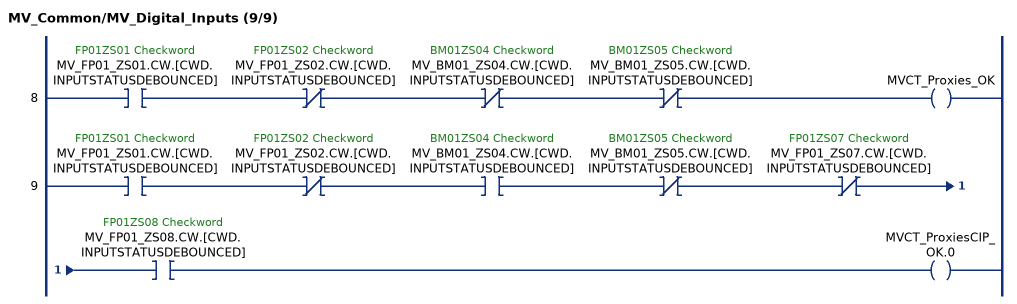
   8: XIC(MV_FP01_ZS01.CW.[CWD.INPUTSTATUSDEBOUNCED])XIO(MV_FP01_ZS02.CW.[CWD.INPUTSTATUSDEBOUNCED])XIO(MV_BM01_ZS04.CW.[CWD.INPUTSTATUSDEBOUNCED])XIO(MV_BM01_ZS05.CW.[CWD.INPUTSTATUSDEBOUNCED])OTE(MVCT_Proxies_OK);
   9: XIC(MV_FP01_ZS01.CW.[CWD.INPUTSTATUSDEBOUNCED])XIO(MV_FP01_ZS02.CW.[CWD.INPUTSTATUSDEBOUNCED])XIC(MV_BM01_ZS04.CW.[CWD.INPUTSTATUSDEBOUNCED])XIO(MV_BM01_ZS05.CW.[CWD.INPUTSTATUSDEBOUNCED])XIO(MV_FP01_ZS07.CW.[CWD.INPUTSTATUSDEBOUNCED])XIC(MV_FP01_ZS08.CW.[CWD.INPUTSTATUSDEBOUNCED])OTE(MVCT_ProxiesCIP_OK.0);
END_ROUTINE

ROUTINE MV_Digital_Outputs   (* ladder *)
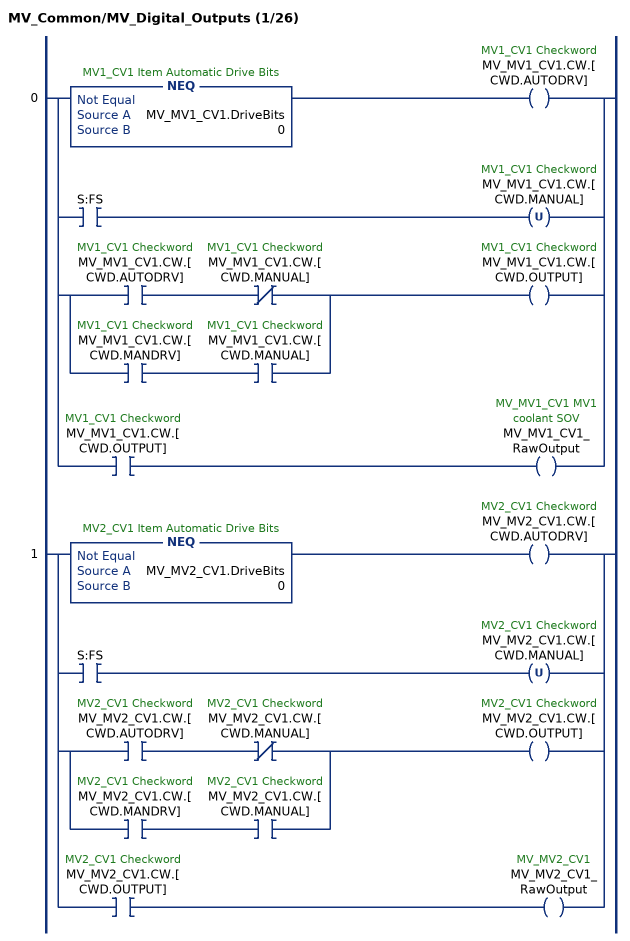
   0: [NEQ(MV_MV1_CV1.DriveBits,0) OTE(MV_MV1_CV1.CW.[CWD.AUTODRV]) ,XIC(S:FS) OTU(MV_MV1_CV1.CW.[CWD.MANUAL]) ,[XIC(MV_MV1_CV1.CW.[CWD.AUTODRV]) XIO(MV_MV1_CV1.CW.[CWD.MANUAL]) ,XIC(MV_MV1_CV1.CW.[CWD.MANDRV]) XIC(MV_MV1_CV1.CW.[CWD.MANUAL]) ] OTE(MV_MV1_CV1.CW.[CWD.OUTPUT]) ,XIC(MV_MV1_CV1.CW.[CWD.OUTPUT]) OTE(MV_MV1_CV1_RawOutput) ];
   1: [NEQ(MV_MV2_CV1.DriveBits,0) OTE(MV_MV2_CV1.CW.[CWD.AUTODRV]) ,XIC(S:FS) OTU(MV_MV2_CV1.CW.[CWD.MANUAL]) ,[XIC(MV_MV2_CV1.CW.[CWD.AUTODRV]) XIO(MV_MV2_CV1.CW.[CWD.MANUAL]) ,XIC(MV_MV2_CV1.CW.[CWD.MANDRV]) XIC(MV_MV2_CV1.CW.[CWD.MANUAL]) ] OTE(MV_MV2_CV1.CW.[CWD.OUTPUT]) ,XIC(MV_MV2_CV1.CW.[CWD.OUTPUT]) OTE(MV_MV2_CV1_RawOutput) ];
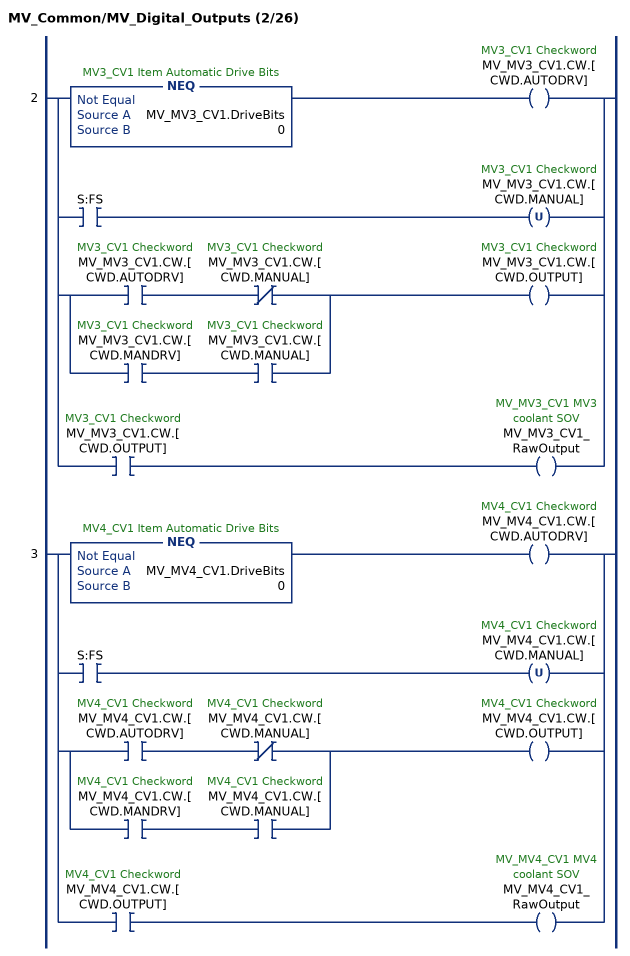
   2: [NEQ(MV_MV3_CV1.DriveBits,0) OTE(MV_MV3_CV1.CW.[CWD.AUTODRV]) ,XIC(S:FS) OTU(MV_MV3_CV1.CW.[CWD.MANUAL]) ,[XIC(MV_MV3_CV1.CW.[CWD.AUTODRV]) XIO(MV_MV3_CV1.CW.[CWD.MANUAL]) ,XIC(MV_MV3_CV1.CW.[CWD.MANDRV]) XIC(MV_MV3_CV1.CW.[CWD.MANUAL]) ] OTE(MV_MV3_CV1.CW.[CWD.OUTPUT]) ,XIC(MV_MV3_CV1.CW.[CWD.OUTPUT]) OTE(MV_MV3_CV1_RawOutput) ];
   3: [NEQ(MV_MV4_CV1.DriveBits,0) OTE(MV_MV4_CV1.CW.[CWD.AUTODRV]) ,XIC(S:FS) OTU(MV_MV4_CV1.CW.[CWD.MANUAL]) ,[XIC(MV_MV4_CV1.CW.[CWD.AUTODRV]) XIO(MV_MV4_CV1.CW.[CWD.MANUAL]) ,XIC(MV_MV4_CV1.CW.[CWD.MANDRV]) XIC(MV_MV4_CV1.CW.[CWD.MANUAL]) ] OTE(MV_MV4_CV1.CW.[CWD.OUTPUT]) ,XIC(MV_MV4_CV1.CW.[CWD.OUTPUT]) OTE(MV_MV4_CV1_RawOutput) ];
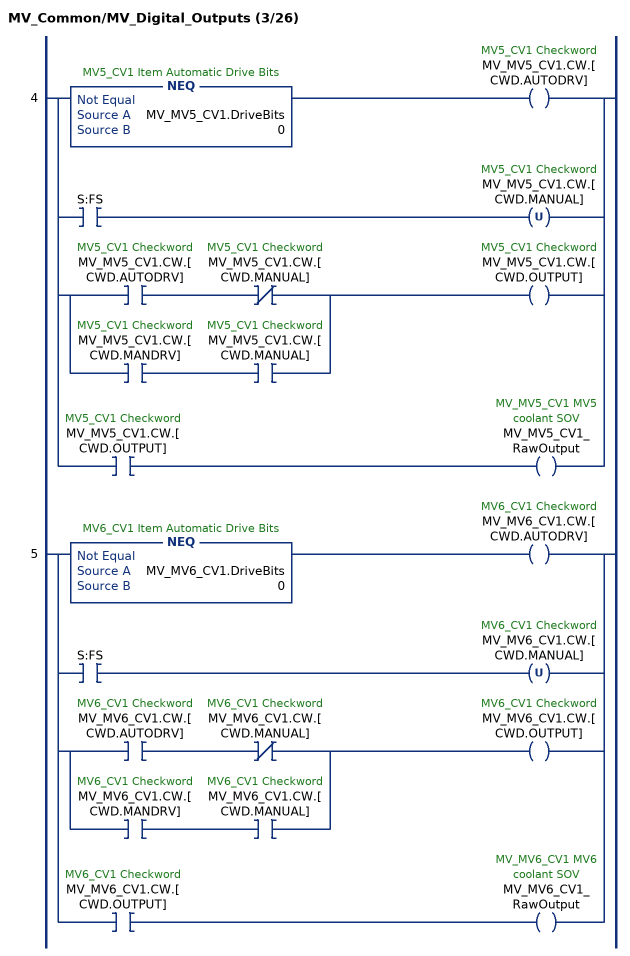
   4: [NEQ(MV_MV5_CV1.DriveBits,0) OTE(MV_MV5_CV1.CW.[CWD.AUTODRV]) ,XIC(S:FS) OTU(MV_MV5_CV1.CW.[CWD.MANUAL]) ,[XIC(MV_MV5_CV1.CW.[CWD.AUTODRV]) XIO(MV_MV5_CV1.CW.[CWD.MANUAL]) ,XIC(MV_MV5_CV1.CW.[CWD.MANDRV]) XIC(MV_MV5_CV1.CW.[CWD.MANUAL]) ] OTE(MV_MV5_CV1.CW.[CWD.OUTPUT]) ,XIC(MV_MV5_CV1.CW.[CWD.OUTPUT]) OTE(MV_MV5_CV1_RawOutput) ];
   5: [NEQ(MV_MV6_CV1.DriveBits,0) OTE(MV_MV6_CV1.CW.[CWD.AUTODRV]) ,XIC(S:FS) OTU(MV_MV6_CV1.CW.[CWD.MANUAL]) ,[XIC(MV_MV6_CV1.CW.[CWD.AUTODRV]) XIO(MV_MV6_CV1.CW.[CWD.MANUAL]) ,XIC(MV_MV6_CV1.CW.[CWD.MANDRV]) XIC(MV_MV6_CV1.CW.[CWD.MANUAL]) ] OTE(MV_MV6_CV1.CW.[CWD.OUTPUT]) ,XIC(MV_MV6_CV1.CW.[CWD.OUTPUT]) OTE(MV_MV6_CV1_RawOutput) ];
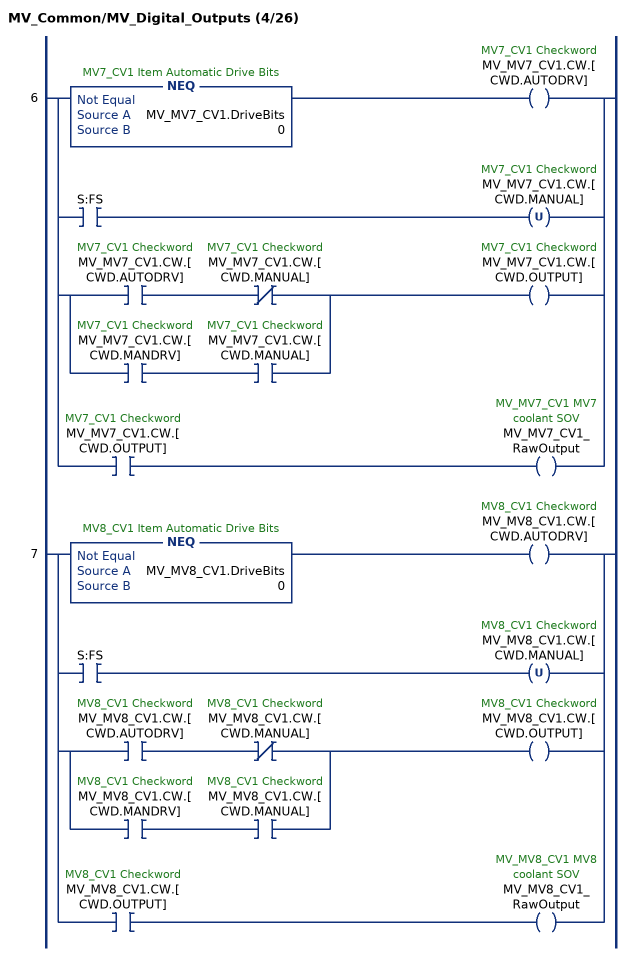
   6: [NEQ(MV_MV7_CV1.DriveBits,0) OTE(MV_MV7_CV1.CW.[CWD.AUTODRV]) ,XIC(S:FS) OTU(MV_MV7_CV1.CW.[CWD.MANUAL]) ,[XIC(MV_MV7_CV1.CW.[CWD.AUTODRV]) XIO(MV_MV7_CV1.CW.[CWD.MANUAL]) ,XIC(MV_MV7_CV1.CW.[CWD.MANDRV]) XIC(MV_MV7_CV1.CW.[CWD.MANUAL]) ] OTE(MV_MV7_CV1.CW.[CWD.OUTPUT]) ,XIC(MV_MV7_CV1.CW.[CWD.OUTPUT]) OTE(MV_MV7_CV1_RawOutput) ];
   7: [NEQ(MV_MV8_CV1.DriveBits,0) OTE(MV_MV8_CV1.CW.[CWD.AUTODRV]) ,XIC(S:FS) OTU(MV_MV8_CV1.CW.[CWD.MANUAL]) ,[XIC(MV_MV8_CV1.CW.[CWD.AUTODRV]) XIO(MV_MV8_CV1.CW.[CWD.MANUAL]) ,XIC(MV_MV8_CV1.CW.[CWD.MANDRV]) XIC(MV_MV8_CV1.CW.[CWD.MANUAL]) ] OTE(MV_MV8_CV1.CW.[CWD.OUTPUT]) ,XIC(MV_MV8_CV1.CW.[CWD.OUTPUT]) OTE(MV_MV8_CV1_RawOutput) ];
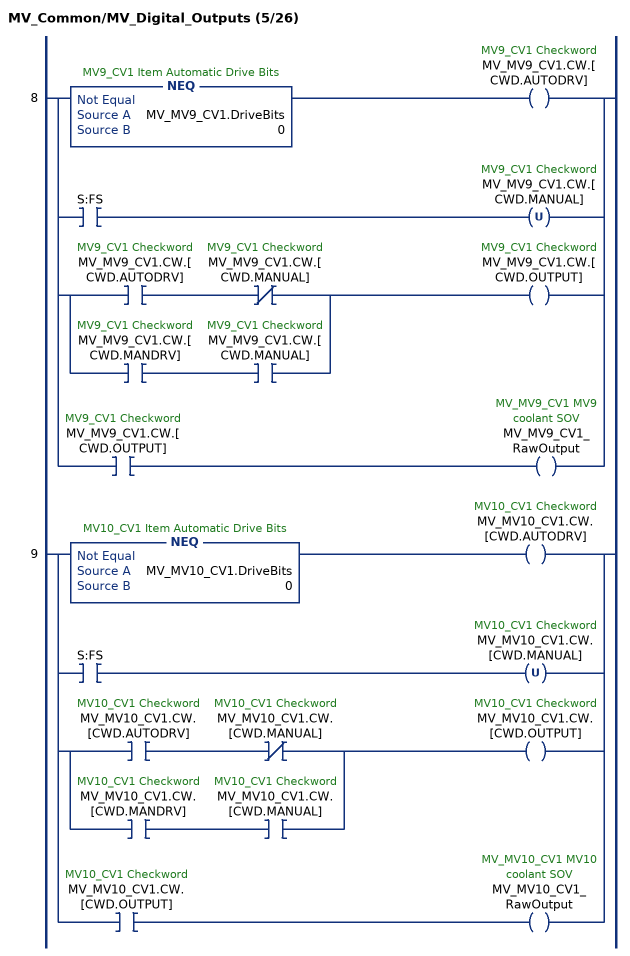
   8: [NEQ(MV_MV9_CV1.DriveBits,0) OTE(MV_MV9_CV1.CW.[CWD.AUTODRV]) ,XIC(S:FS) OTU(MV_MV9_CV1.CW.[CWD.MANUAL]) ,[XIC(MV_MV9_CV1.CW.[CWD.AUTODRV]) XIO(MV_MV9_CV1.CW.[CWD.MANUAL]) ,XIC(MV_MV9_CV1.CW.[CWD.MANDRV]) XIC(MV_MV9_CV1.CW.[CWD.MANUAL]) ] OTE(MV_MV9_CV1.CW.[CWD.OUTPUT]) ,XIC(MV_MV9_CV1.CW.[CWD.OUTPUT]) OTE(MV_MV9_CV1_RawOutput) ];
   9: [NEQ(MV_MV10_CV1.DriveBits,0) OTE(MV_MV10_CV1.CW.[CWD.AUTODRV]) ,XIC(S:FS) OTU(MV_MV10_CV1.CW.[CWD.MANUAL]) ,[XIC(MV_MV10_CV1.CW.[CWD.AUTODRV]) XIO(MV_MV10_CV1.CW.[CWD.MANUAL]) ,XIC(MV_MV10_CV1.CW.[CWD.MANDRV]) XIC(MV_MV10_CV1.CW.[CWD.MANUAL]) ] OTE(MV_MV10_CV1.CW.[CWD.OUTPUT]) ,XIC(MV_MV10_CV1.CW.[CWD.OUTPUT]) OTE(MV_MV10_CV1_RawOutput) ];
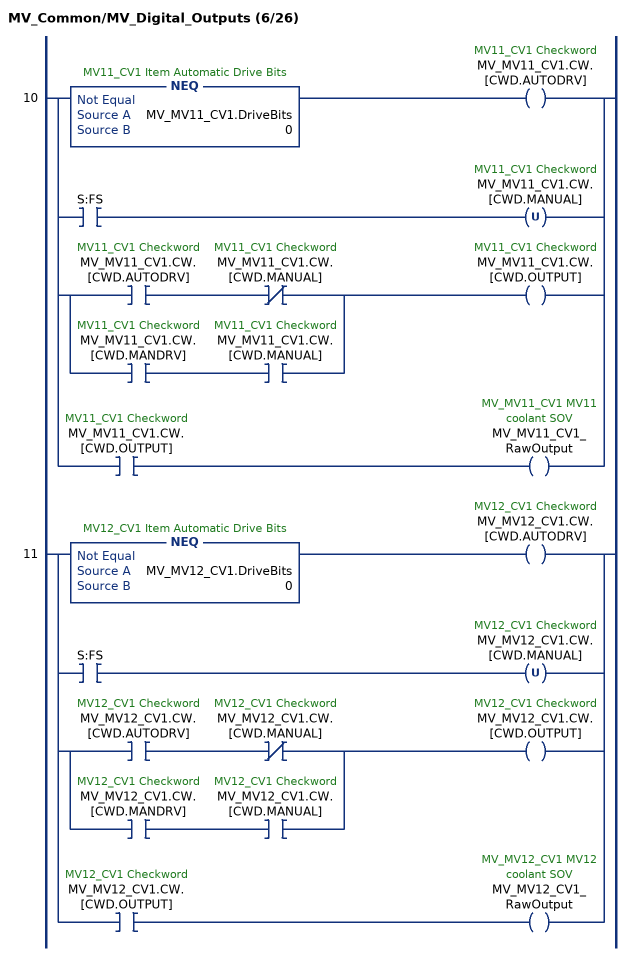
   10: [NEQ(MV_MV11_CV1.DriveBits,0) OTE(MV_MV11_CV1.CW.[CWD.AUTODRV]) ,XIC(S:FS) OTU(MV_MV11_CV1.CW.[CWD.MANUAL]) ,[XIC(MV_MV11_CV1.CW.[CWD.AUTODRV]) XIO(MV_MV11_CV1.CW.[CWD.MANUAL]) ,XIC(MV_MV11_CV1.CW.[CWD.MANDRV]) XIC(MV_MV11_CV1.CW.[CWD.MANUAL]) ] OTE(MV_MV11_CV1.CW.[CWD.OUTPUT]) ,XIC(MV_MV11_CV1.CW.[CWD.OUTPUT]) OTE(MV_MV11_CV1_RawOutput) ];
   11: [NEQ(MV_MV12_CV1.DriveBits,0) OTE(MV_MV12_CV1.CW.[CWD.AUTODRV]) ,XIC(S:FS) OTU(MV_MV12_CV1.CW.[CWD.MANUAL]) ,[XIC(MV_MV12_CV1.CW.[CWD.AUTODRV]) XIO(MV_MV12_CV1.CW.[CWD.MANUAL]) ,XIC(MV_MV12_CV1.CW.[CWD.MANDRV]) XIC(MV_MV12_CV1.CW.[CWD.MANUAL]) ] OTE(MV_MV12_CV1.CW.[CWD.OUTPUT]) ,XIC(MV_MV12_CV1.CW.[CWD.OUTPUT]) OTE(MV_MV12_CV1_RawOutput) ];
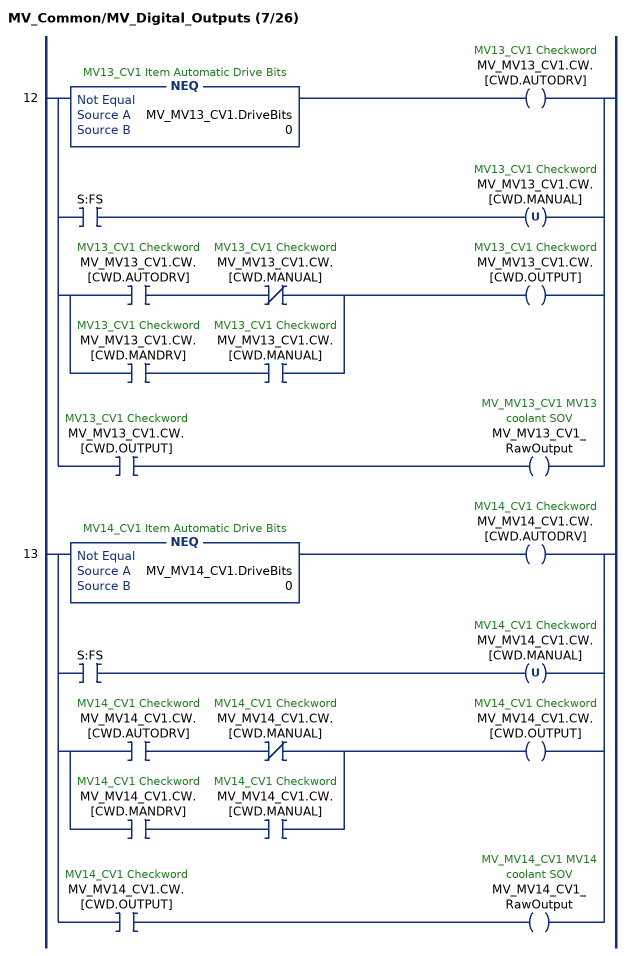
   12: [NEQ(MV_MV13_CV1.DriveBits,0) OTE(MV_MV13_CV1.CW.[CWD.AUTODRV]) ,XIC(S:FS) OTU(MV_MV13_CV1.CW.[CWD.MANUAL]) ,[XIC(MV_MV13_CV1.CW.[CWD.AUTODRV]) XIO(MV_MV13_CV1.CW.[CWD.MANUAL]) ,XIC(MV_MV13_CV1.CW.[CWD.MANDRV]) XIC(MV_MV13_CV1.CW.[CWD.MANUAL]) ] OTE(MV_MV13_CV1.CW.[CWD.OUTPUT]) ,XIC(MV_MV13_CV1.CW.[CWD.OUTPUT]) OTE(MV_MV13_CV1_RawOutput) ];
   13: [NEQ(MV_MV14_CV1.DriveBits,0) OTE(MV_MV14_CV1.CW.[CWD.AUTODRV]) ,XIC(S:FS) OTU(MV_MV14_CV1.CW.[CWD.MANUAL]) ,[XIC(MV_MV14_CV1.CW.[CWD.AUTODRV]) XIO(MV_MV14_CV1.CW.[CWD.MANUAL]) ,XIC(MV_MV14_CV1.CW.[CWD.MANDRV]) XIC(MV_MV14_CV1.CW.[CWD.MANUAL]) ] OTE(MV_MV14_CV1.CW.[CWD.OUTPUT]) ,XIC(MV_MV14_CV1.CW.[CWD.OUTPUT]) OTE(MV_MV14_CV1_RawOutput) ];
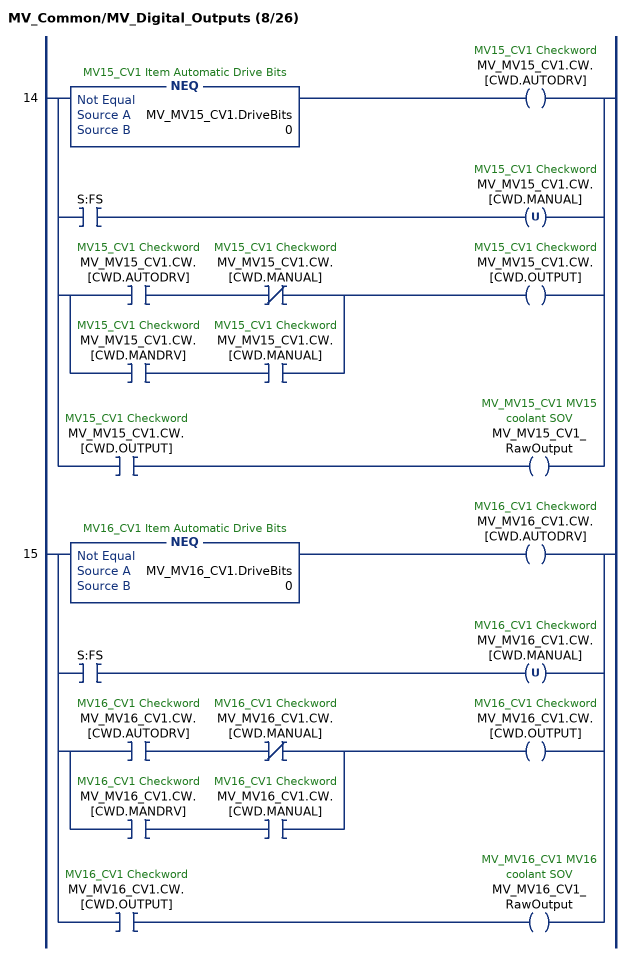
   14: [NEQ(MV_MV15_CV1.DriveBits,0) OTE(MV_MV15_CV1.CW.[CWD.AUTODRV]) ,XIC(S:FS) OTU(MV_MV15_CV1.CW.[CWD.MANUAL]) ,[XIC(MV_MV15_CV1.CW.[CWD.AUTODRV]) XIO(MV_MV15_CV1.CW.[CWD.MANUAL]) ,XIC(MV_MV15_CV1.CW.[CWD.MANDRV]) XIC(MV_MV15_CV1.CW.[CWD.MANUAL]) ] OTE(MV_MV15_CV1.CW.[CWD.OUTPUT]) ,XIC(MV_MV15_CV1.CW.[CWD.OUTPUT]) OTE(MV_MV15_CV1_RawOutput) ];
   15: [NEQ(MV_MV16_CV1.DriveBits,0) OTE(MV_MV16_CV1.CW.[CWD.AUTODRV]) ,XIC(S:FS) OTU(MV_MV16_CV1.CW.[CWD.MANUAL]) ,[XIC(MV_MV16_CV1.CW.[CWD.AUTODRV]) XIO(MV_MV16_CV1.CW.[CWD.MANUAL]) ,XIC(MV_MV16_CV1.CW.[CWD.MANDRV]) XIC(MV_MV16_CV1.CW.[CWD.MANUAL]) ] OTE(MV_MV16_CV1.CW.[CWD.OUTPUT]) ,XIC(MV_MV16_CV1.CW.[CWD.OUTPUT]) OTE(MV_MV16_CV1_RawOutput) ];
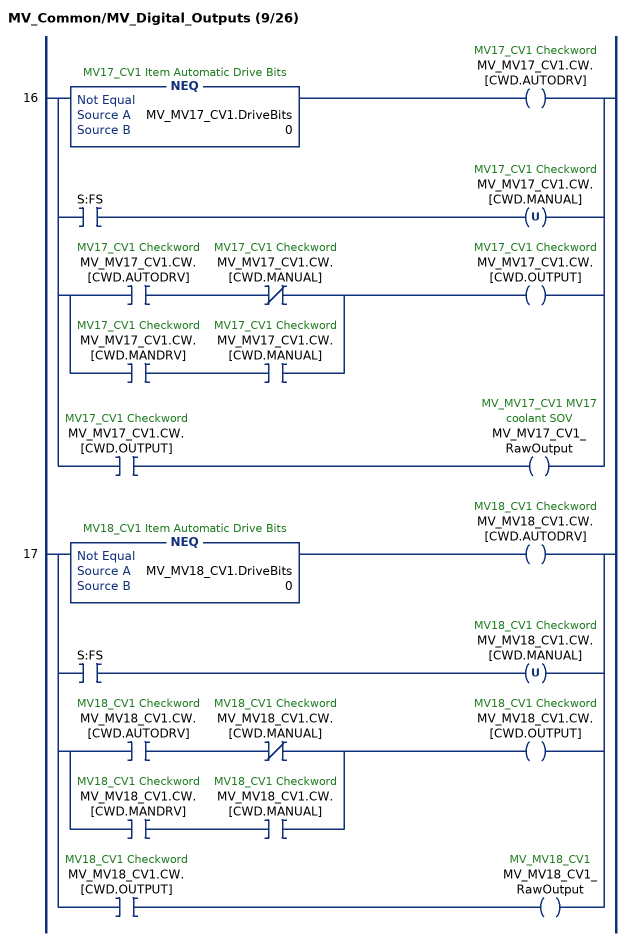
   16: [NEQ(MV_MV17_CV1.DriveBits,0) OTE(MV_MV17_CV1.CW.[CWD.AUTODRV]) ,XIC(S:FS) OTU(MV_MV17_CV1.CW.[CWD.MANUAL]) ,[XIC(MV_MV17_CV1.CW.[CWD.AUTODRV]) XIO(MV_MV17_CV1.CW.[CWD.MANUAL]) ,XIC(MV_MV17_CV1.CW.[CWD.MANDRV]) XIC(MV_MV17_CV1.CW.[CWD.MANUAL]) ] OTE(MV_MV17_CV1.CW.[CWD.OUTPUT]) ,XIC(MV_MV17_CV1.CW.[CWD.OUTPUT]) OTE(MV_MV17_CV1_RawOutput) ];
   17: [NEQ(MV_MV18_CV1.DriveBits,0) OTE(MV_MV18_CV1.CW.[CWD.AUTODRV]) ,XIC(S:FS) OTU(MV_MV18_CV1.CW.[CWD.MANUAL]) ,[XIC(MV_MV18_CV1.CW.[CWD.AUTODRV]) XIO(MV_MV18_CV1.CW.[CWD.MANUAL]) ,XIC(MV_MV18_CV1.CW.[CWD.MANDRV]) XIC(MV_MV18_CV1.CW.[CWD.MANUAL]) ] OTE(MV_MV18_CV1.CW.[CWD.OUTPUT]) ,XIC(MV_MV18_CV1.CW.[CWD.OUTPUT]) OTE(MV_MV18_CV1_RawOutput) ];
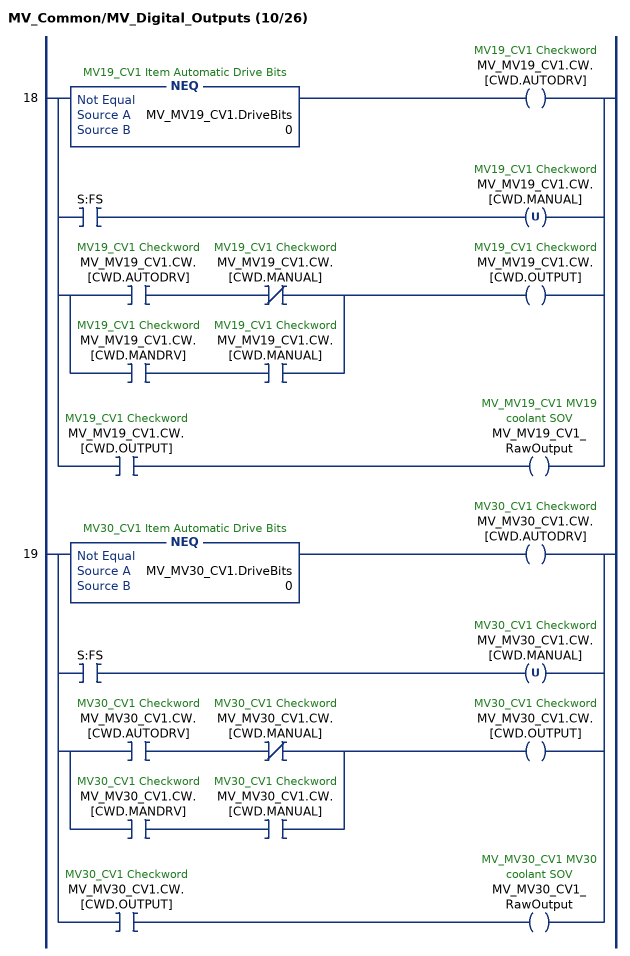
   18: [NEQ(MV_MV19_CV1.DriveBits,0) OTE(MV_MV19_CV1.CW.[CWD.AUTODRV]) ,XIC(S:FS) OTU(MV_MV19_CV1.CW.[CWD.MANUAL]) ,[XIC(MV_MV19_CV1.CW.[CWD.AUTODRV]) XIO(MV_MV19_CV1.CW.[CWD.MANUAL]) ,XIC(MV_MV19_CV1.CW.[CWD.MANDRV]) XIC(MV_MV19_CV1.CW.[CWD.MANUAL]) ] OTE(MV_MV19_CV1.CW.[CWD.OUTPUT]) ,XIC(MV_MV19_CV1.CW.[CWD.OUTPUT]) OTE(MV_MV19_CV1_RawOutput) ];
   19: [NEQ(MV_MV30_CV1.DriveBits,0) OTE(MV_MV30_CV1.CW.[CWD.AUTODRV]) ,XIC(S:FS) OTU(MV_MV30_CV1.CW.[CWD.MANUAL]) ,[XIC(MV_MV30_CV1.CW.[CWD.AUTODRV]) XIO(MV_MV30_CV1.CW.[CWD.MANUAL]) ,XIC(MV_MV30_CV1.CW.[CWD.MANDRV]) XIC(MV_MV30_CV1.CW.[CWD.MANUAL]) ] OTE(MV_MV30_CV1.CW.[CWD.OUTPUT]) ,XIC(MV_MV30_CV1.CW.[CWD.OUTPUT]) OTE(MV_MV30_CV1_RawOutput) ];
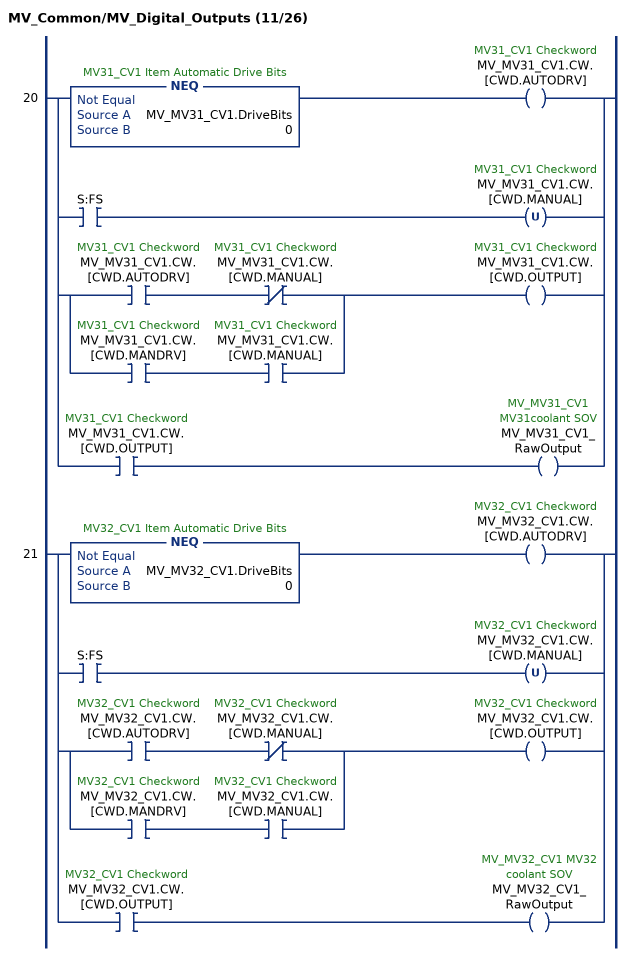
   20: [NEQ(MV_MV31_CV1.DriveBits,0) OTE(MV_MV31_CV1.CW.[CWD.AUTODRV]) ,XIC(S:FS) OTU(MV_MV31_CV1.CW.[CWD.MANUAL]) ,[XIC(MV_MV31_CV1.CW.[CWD.AUTODRV]) XIO(MV_MV31_CV1.CW.[CWD.MANUAL]) ,XIC(MV_MV31_CV1.CW.[CWD.MANDRV]) XIC(MV_MV31_CV1.CW.[CWD.MANUAL]) ] OTE(MV_MV31_CV1.CW.[CWD.OUTPUT]) ,XIC(MV_MV31_CV1.CW.[CWD.OUTPUT]) OTE(MV_MV31_CV1_RawOutput) ];
   21: [NEQ(MV_MV32_CV1.DriveBits,0) OTE(MV_MV32_CV1.CW.[CWD.AUTODRV]) ,XIC(S:FS) OTU(MV_MV32_CV1.CW.[CWD.MANUAL]) ,[XIC(MV_MV32_CV1.CW.[CWD.AUTODRV]) XIO(MV_MV32_CV1.CW.[CWD.MANUAL]) ,XIC(MV_MV32_CV1.CW.[CWD.MANDRV]) XIC(MV_MV32_CV1.CW.[CWD.MANUAL]) ] OTE(MV_MV32_CV1.CW.[CWD.OUTPUT]) ,XIC(MV_MV32_CV1.CW.[CWD.OUTPUT]) OTE(MV_MV32_CV1_RawOutput) ];
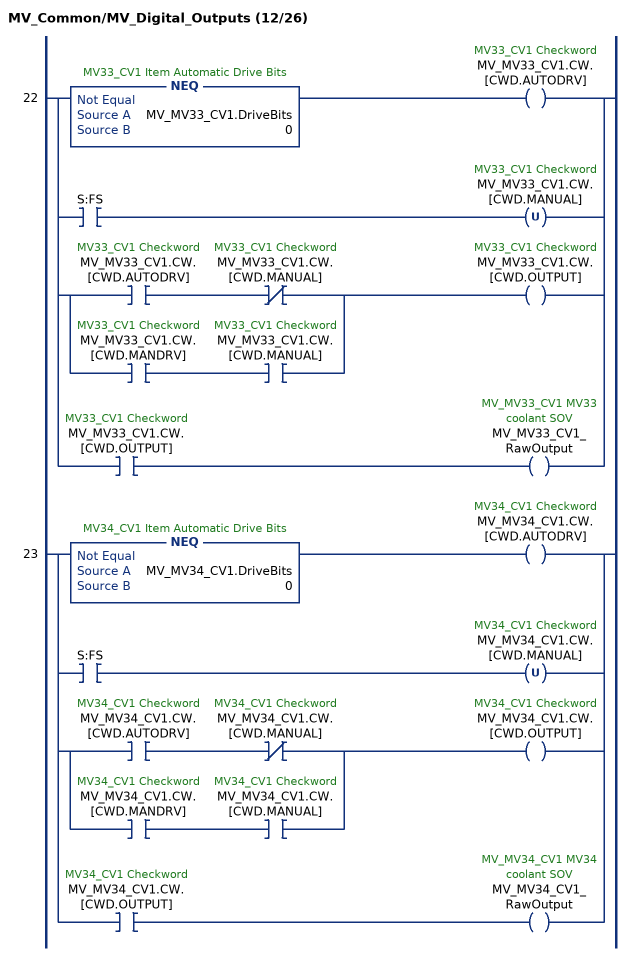
   22: [NEQ(MV_MV33_CV1.DriveBits,0) OTE(MV_MV33_CV1.CW.[CWD.AUTODRV]) ,XIC(S:FS) OTU(MV_MV33_CV1.CW.[CWD.MANUAL]) ,[XIC(MV_MV33_CV1.CW.[CWD.AUTODRV]) XIO(MV_MV33_CV1.CW.[CWD.MANUAL]) ,XIC(MV_MV33_CV1.CW.[CWD.MANDRV]) XIC(MV_MV33_CV1.CW.[CWD.MANUAL]) ] OTE(MV_MV33_CV1.CW.[CWD.OUTPUT]) ,XIC(MV_MV33_CV1.CW.[CWD.OUTPUT]) OTE(MV_MV33_CV1_RawOutput) ];
   23: [NEQ(MV_MV34_CV1.DriveBits,0) OTE(MV_MV34_CV1.CW.[CWD.AUTODRV]) ,XIC(S:FS) OTU(MV_MV34_CV1.CW.[CWD.MANUAL]) ,[XIC(MV_MV34_CV1.CW.[CWD.AUTODRV]) XIO(MV_MV34_CV1.CW.[CWD.MANUAL]) ,XIC(MV_MV34_CV1.CW.[CWD.MANDRV]) XIC(MV_MV34_CV1.CW.[CWD.MANUAL]) ] OTE(MV_MV34_CV1.CW.[CWD.OUTPUT]) ,XIC(MV_MV34_CV1.CW.[CWD.OUTPUT]) OTE(MV_MV34_CV1_RawOutput) ];
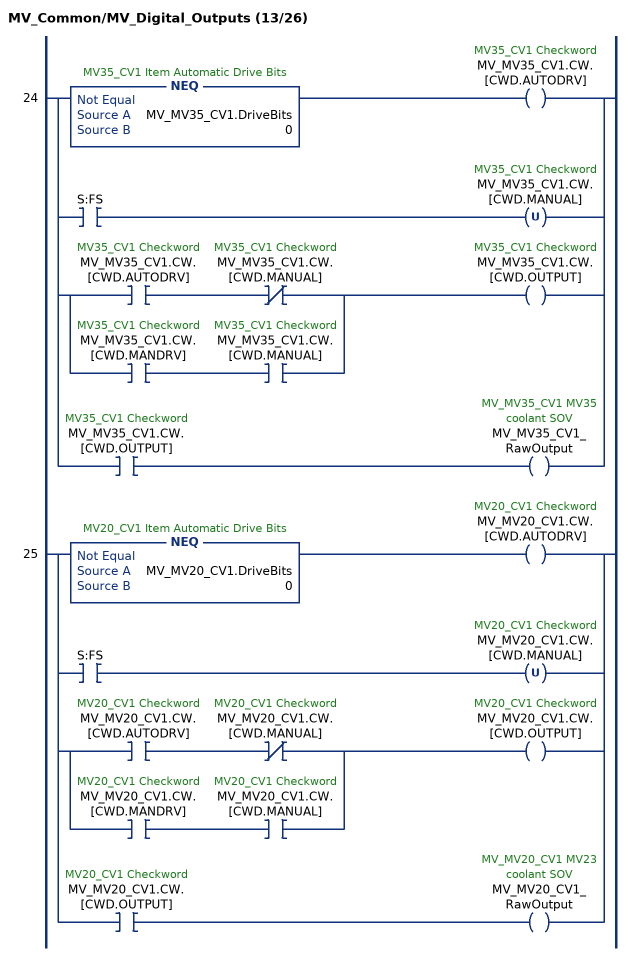
   24: [NEQ(MV_MV35_CV1.DriveBits,0) OTE(MV_MV35_CV1.CW.[CWD.AUTODRV]) ,XIC(S:FS) OTU(MV_MV35_CV1.CW.[CWD.MANUAL]) ,[XIC(MV_MV35_CV1.CW.[CWD.AUTODRV]) XIO(MV_MV35_CV1.CW.[CWD.MANUAL]) ,XIC(MV_MV35_CV1.CW.[CWD.MANDRV]) XIC(MV_MV35_CV1.CW.[CWD.MANUAL]) ] OTE(MV_MV35_CV1.CW.[CWD.OUTPUT]) ,XIC(MV_MV35_CV1.CW.[CWD.OUTPUT]) OTE(MV_MV35_CV1_RawOutput) ];
   25: [NEQ(MV_MV20_CV1.DriveBits,0) OTE(MV_MV20_CV1.CW.[CWD.AUTODRV]) ,XIC(S:FS) OTU(MV_MV20_CV1.CW.[CWD.MANUAL]) ,[XIC(MV_MV20_CV1.CW.[CWD.AUTODRV]) XIO(MV_MV20_CV1.CW.[CWD.MANUAL]) ,XIC(MV_MV20_CV1.CW.[CWD.MANDRV]) XIC(MV_MV20_CV1.CW.[CWD.MANUAL]) ] OTE(MV_MV20_CV1.CW.[CWD.OUTPUT]) ,XIC(MV_MV20_CV1.CW.[CWD.OUTPUT]) OTE(MV_MV20_CV1_RawOutput) ];
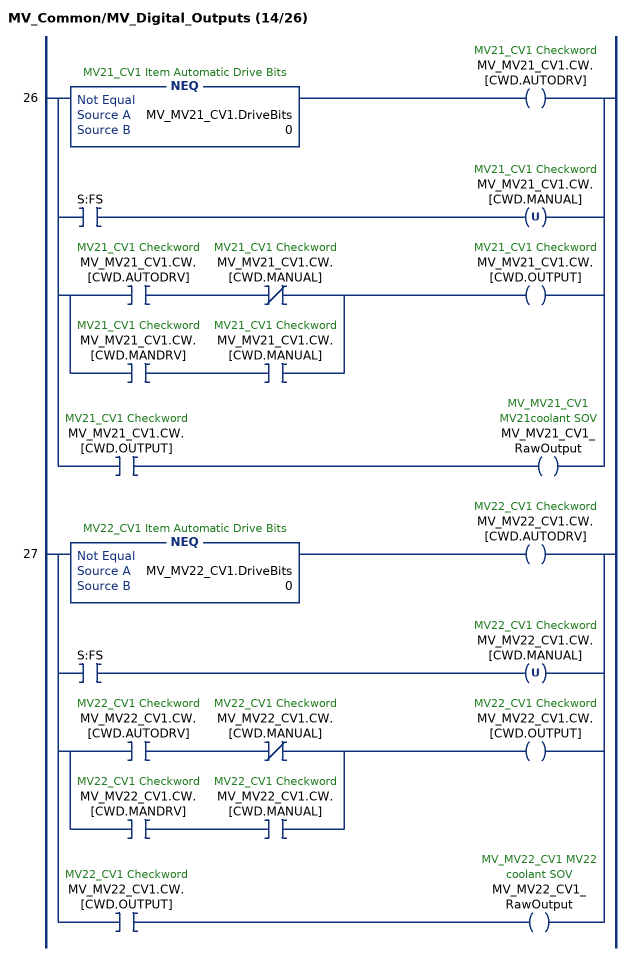
   26: [NEQ(MV_MV21_CV1.DriveBits,0) OTE(MV_MV21_CV1.CW.[CWD.AUTODRV]) ,XIC(S:FS) OTU(MV_MV21_CV1.CW.[CWD.MANUAL]) ,[XIC(MV_MV21_CV1.CW.[CWD.AUTODRV]) XIO(MV_MV21_CV1.CW.[CWD.MANUAL]) ,XIC(MV_MV21_CV1.CW.[CWD.MANDRV]) XIC(MV_MV21_CV1.CW.[CWD.MANUAL]) ] OTE(MV_MV21_CV1.CW.[CWD.OUTPUT]) ,XIC(MV_MV21_CV1.CW.[CWD.OUTPUT]) OTE(MV_MV21_CV1_RawOutput) ];
   27: [NEQ(MV_MV22_CV1.DriveBits,0) OTE(MV_MV22_CV1.CW.[CWD.AUTODRV]) ,XIC(S:FS) OTU(MV_MV22_CV1.CW.[CWD.MANUAL]) ,[XIC(MV_MV22_CV1.CW.[CWD.AUTODRV]) XIO(MV_MV22_CV1.CW.[CWD.MANUAL]) ,XIC(MV_MV22_CV1.CW.[CWD.MANDRV]) XIC(MV_MV22_CV1.CW.[CWD.MANUAL]) ] OTE(MV_MV22_CV1.CW.[CWD.OUTPUT]) ,XIC(MV_MV22_CV1.CW.[CWD.OUTPUT]) OTE(MV_MV22_CV1_RawOutput) ];
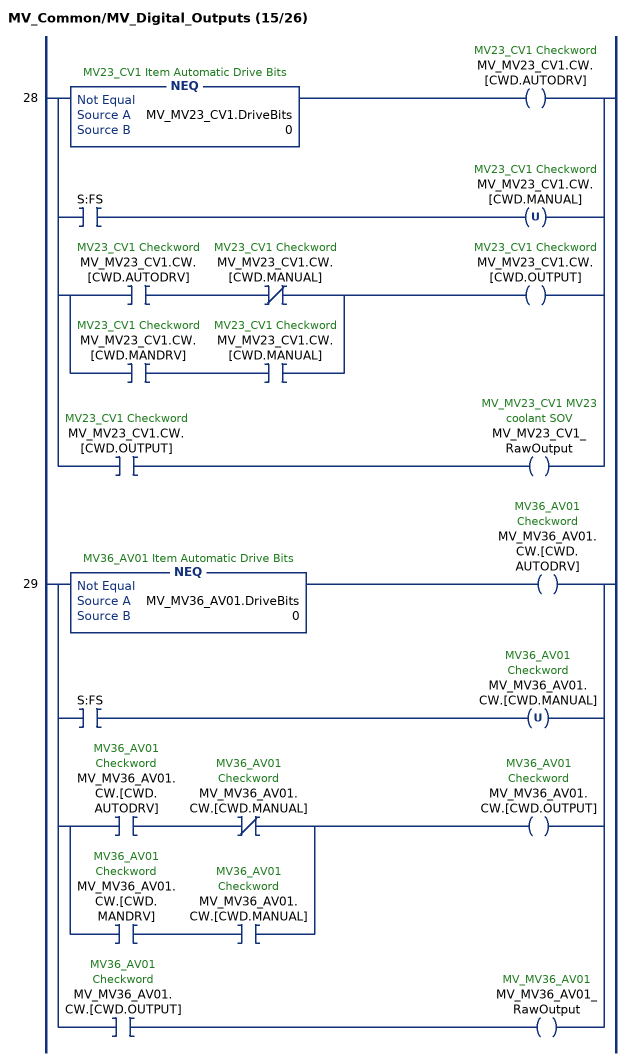
   28: [NEQ(MV_MV23_CV1.DriveBits,0) OTE(MV_MV23_CV1.CW.[CWD.AUTODRV]) ,XIC(S:FS) OTU(MV_MV23_CV1.CW.[CWD.MANUAL]) ,[XIC(MV_MV23_CV1.CW.[CWD.AUTODRV]) XIO(MV_MV23_CV1.CW.[CWD.MANUAL]) ,XIC(MV_MV23_CV1.CW.[CWD.MANDRV]) XIC(MV_MV23_CV1.CW.[CWD.MANUAL]) ] OTE(MV_MV23_CV1.CW.[CWD.OUTPUT]) ,XIC(MV_MV23_CV1.CW.[CWD.OUTPUT]) OTE(MV_MV23_CV1_RawOutput) ];
   29: [NEQ(MV_MV36_AV01.DriveBits,0) OTE(MV_MV36_AV01.CW.[CWD.AUTODRV]) ,XIC(S:FS) OTU(MV_MV36_AV01.CW.[CWD.MANUAL]) ,[XIC(MV_MV36_AV01.CW.[CWD.AUTODRV]) XIO(MV_MV36_AV01.CW.[CWD.MANUAL]) ,XIC(MV_MV36_AV01.CW.[CWD.MANDRV]) XIC(MV_MV36_AV01.CW.[CWD.MANUAL]) ] OTE(MV_MV36_AV01.CW.[CWD.OUTPUT]) ,XIC(MV_MV36_AV01.CW.[CWD.OUTPUT]) OTE(MV_MV36_AV01_RawOutput) ];
